
screen "Root screen" 800x480, template "Main"
   Rectangle "Rectangle_1" at 7,7 size 265x142
      Appearance <- "Comm_1_DB_Warning"
   GraphicView "Graphic view_4" at 169,29 size 84x118; Picture "h2o_1"
   GraphicView "Graphic view_2" at 89,29 size 84x118; Picture "h2o_1"
   Bar "Bar_1" at 229,7 size 43x142; Unit %; MinimumValue 0; MaximumValue 100
      ProcessValue <- "Comm_1_DB_Level"
   GraphicView "Graphic view_1" at 9,29 size 84x118; Picture "h2o_1"
   GraphicIOField "Graphic I/O field_7" at 101,119 size 76x24; PictureList "L_1"
      ProcessValue <- "Comm_1_DB_Mix_2_Status"
   GraphicIOField "Graphic I/O field_8" at 191,119 size 76x24; PictureList "L_1"
      ProcessValue <- "Comm_1_DB_Mix_3_Status"
   GraphicIOField "Graphic I/O field_6" at 12,119 size 76x24; PictureList "L_1"
      ProcessValue <- "Comm_1_DB_Mix_1_Status"
   TextField "Text field_4" at 447,6 size 223x27; Text 'мастер шкаф дозации'
   TextField "Text field_5" at 447,27 size 227x72; Text 'PolyMix'
   Button "Button_8" at 543,238 size 175x60; TextOff 'Авто'
      on Click: SetBit("Logick_DB_Start")
      Appearance <- "Logick_DB_Start"
   Button "Button_9" at 543,326 size 175x60; TextOff 'Стоп'
      on Click: ResetBit("Logick_DB_Start")
   Button "Button_10" at 543,415 size 175x60; TextOff 'Ручной'; Authorization "Operator"
      on Click: InvertBit("Logick_DB_Hand")
      Appearance <- "Logick_DB_Hand"
   Group "Group" at 7,7 size 265x142; Picture "h2o_1"; PictureList "L_1"
   Group "Group_1" at 7,160 size 265x142; Picture "h2o_1"; PictureList "L_1"
   GraphicIOField "Graphic I/O field_4" at 7,312 size 90x90; PictureList "Pump"
      ProcessValue <- "Motors_DB_M1_Status"
   GraphicIOField "Graphic I/O field_5" at 221,312 size 90x90; PictureList "Pump"
      ProcessValue <- "Motors_DB_M2_Status"
   GraphicIOField "Graphic I/O field_9" at 439,312 size 90x90; PictureList "Pump"
      ProcessValue <- "Motors_DB_M3_Status"
   Button "Button_7" at 7,402 size 90x22; TextOff 'Активен'; TextList "Hand"
      on Click: InvertBit("Logick_DB_Use_M1")
      ProcessValue <- "Motors_DB_M1_CMD_Hand"
      Appearance <- "Logick_DB_Use_M1"
   Button "Button_1" at 439,402 size 90x22; TextOff 'Активен'; TextList "Hand"
      on Click: InvertBit("Logick_DB_Use_M3")
      ProcessValue <- "Motors_DB_M1_CMD_Hand"
      Appearance <- "Logick_DB_Use_M3"
   Button "Button_2" at 221,402 size 90x22; TextOff 'Резерв М1'; TextList "Hand"
      on Click: SetBit("Logick_DB_Res_M1"); ResetBit("Logick_DB_Res_M3")
      ProcessValue <- "Motors_DB_M1_CMD_Hand"
      Appearance <- "Logick_DB_Res_M1"
   Button "Button_3" at 221,429 size 90x22; TextOff 'Резерв М3'; TextList "Hand"
      on Click: SetBit("Logick_DB_Res_M3"); ResetBit("Logick_DB_Res_M1")
      ProcessValue <- "Motors_DB_M1_CMD_Hand"
      Appearance <- "Logick_DB_Res_M3"
   Button "Button_4" at 221,457 size 90x22; TextOff 'Стоп'; TextList "Hand"
      on Click: ResetBit("Logick_DB_Res_M3"); ResetBit("Logick_DB_Res_M1")
      ProcessValue <- "Motors_DB_M1_CMD_Hand"
   GraphicView "Graphic view_7" at 275,7 size 156x149; Picture "Graphic_9"
   GraphicView "Graphic view_8" at 276,160 size 156x149; Picture "Graphic_9"
   IOField "I/O field_17" at 308,18 size 98x30; FormatPattern 99999.99
      ProcessValue <- "Statistics_DB_Mass_1"
      Appearance <- "DIx_DB_Mass_1_Signal"
   TextField "Text field_1" at 345,43 size 25x27; Text 'кг'
   IOField "I/O field_1" at 308,109 size 98x30; FormatPattern 99999.99
      ProcessValue <- "Statistics_DB_Today_1"
      Appearance <- "DIx_DB_Mass_1_Signal"
   TextField "Text field_2" at 315,83 size 85x27; Text 'за день:'
   IOField "I/O field_2" at 308,171 size 98x30; FormatPattern 99999.99
      ProcessValue <- "Statistics_DB_Mass_2"
      Appearance <- "DIx_DB_Mass_2_Signal"
   TextField "Text field_3" at 345,196 size 25x27; Text 'кг'
   IOField "I/O field_3" at 308,262 size 98x30; FormatPattern 99999.99
      ProcessValue <- "Statistics_DB_Today_2"
      Appearance <- "DIx_DB_Mass_2_Signal"
   TextField "Text field_6" at 315,236 size 85x27; Text 'за день:'
   IOField "I/O field_4" at 7,432 size 92x30; FormatPattern 9999.99
      Appearance <- "Logick_DB_Low_REQ"
      ProcessValue <- "AIx_DB_Flow_1_Result"
   TextField "Text field_7" at 33,453 size 40x27; Text 'л/ч'
   IOField "I/O field_5" at 438,432 size 92x30; FormatPattern 9999.99
      Appearance <- "Logick_DB_Low_REQ"
      ProcessValue <- "AIx_DB_Flow_2_Result"
   TextField "Text field_8" at 464,453 size 40x27; Text 'л/ч'
   Button "Button_5" at 128,362 size 60x60; TextOff 'Text'; PictureOff "table"
      on Click: ActivateScreen("Point_1", 0)
   Button "Button_6" at 348,362 size 60x60; TextOff 'Text'; PictureOff "table"
      on Click: ActivateScreen("Point_2", 0)
   TextField "Text field_9" at 347,304 size 60x27; Text 'Доза:'
   TextField "Text field_11" at 32,339 size 34x27; Text 'М1'
   TextField "Text field_12" at 247,338 size 34x27; Text 'М2'
   TextField "Text field_13" at 465,337 size 34x27; Text 'М3'
   IOField "I/O field_7" at 119,328 size 77x30; FormatPattern 999.99
      ProcessValue <- "Logick_DB_D_1"
      Visibility <- "Logick_DB_Fix_1"
   TextField "Text field_14" at 128,303 size 60x27; Text 'Доза:'
   Button "Button_12" at 118,424 size 80x25; TextOff 'Text'; Authorization "Operator"; PictureList "ON_OFF"
      on Click: InvertBit("Logick_DB_Fix_1")
      ProcessValue <- "Logick_DB_Fix_1"
   IOField "I/O field_8" at 119,328 size 77x30; Authorization "Operator"; FormatPattern 999.99
      ProcessValue <- "Logick_DB_Fix_D_1"
      Visibility <- "Logick_DB_Fix_1"
   IOField "I/O field_6" at 339,329 size 77x30; FormatPattern 999.99
      Visibility <- "Logick_DB_Fix_2"
      ProcessValue <- "Logick_DB_D_2"
   Button "Button_11" at 339,424 size 80x25; TextOff 'Text'; PictureList "ON_OFF"; Authorization "Operator"
      on Click: InvertBit("Logick_DB_Fix_2")
      ProcessValue <- "Logick_DB_Fix_2"
   IOField "I/O field_9" at 339,329 size 77x30; Authorization "Operator"; FormatPattern 999.99
      Visibility <- "Logick_DB_Fix_2"
      ProcessValue <- "Logick_DB_Fix_D_2"
   Button "Button_13" at 8,312 size 86x86; TextOff 'Text'
      on Click: InvertBit("Motors_DB_M1_CMD_Start_M")
   Button "Button_14" at 223,312 size 86x86; TextOff 'Text'
      on Click: InvertBit("Motors_DB_M2_CMD_Start_M")
   Button "Button_15" at 441,312 size 86x86; TextOff 'Text'
      on Click: InvertBit("Motors_DB_M3_CMD_Start_M")
   TextField "Text field_16" at 447,99 size 220x27; Text 'Производительность:'
   TextField "Text field_17" at 447,127 size 112x27; Text 'Дозатор 1:'
   TextField "Text field_18" at 447,163 size 112x27; Text 'Дозатор 2:'
   TextField "Text field_19" at 447,200 size 112x27; Text 'Дозатор 3:'
   IOField "I/O field_10" at 558,127 size 77x30; Authorization "Operator"; FormatPattern 9999
      ProcessValue <- "AOx_DB_M1_SP_SP_M"
      Appearance <- "AOx_DB_M1_SP_CMD_Hand"
   IOField "I/O field_11" at 558,162 size 77x30; Authorization "Operator"; FormatPattern 9999
      Appearance <- "AOx_DB_M2_SP_CMD_Hand"
      ProcessValue <- "AOx_DB_M2_SP_SP_M"
   IOField "I/O field_12" at 558,197 size 77x30; Authorization "Operator"; FormatPattern 9999
      Appearance <- "AOx_DB_M3_SP_CMD_Hand"
      ProcessValue <- "AOx_DB_M3_SP_SP_M"
   IOField "I/O field_13" at 339,448 size 80x30; FormatPattern 999.99
      ProcessValue <- "AIx_DB_Trans_2_Result"
   IOField "I/O field_14" at 118,448 size 80x30; FormatPattern 999.99
      ProcessValue <- "AIx_DB_Trans_1_Result"
   Button "Button_16" at 278,6 size 149x139; TextOff 'Text'
      on Click: ActivateScreen("Mass_1", 0)
   Button "Button_17" at 280,159 size 149x139; TextOff 'Text'
      on Click: ActivateScreen("Mass_2", 0)
   GraphicView "Graphic view_9" at 447,236 size 30x30; Picture "heat"
      Appearance <- "DIx_DB_Heat_1_Signal"
   GraphicView "Graphic view_10" at 492,236 size 30x30; Picture "heat"
      Appearance <- "DIx_DB_Heat_2_Signal"
   GraphicView "Graphic view_11" at 448,274 size 30x30; Picture "heat"
      Appearance <- "DIx_DB_Heat_3_Signal"
   GraphicView "Graphic view_12" at 492,274 size 30x30; Picture "heat"
      Appearance <- "DIx_DB_Heat_4_Signal"
   IOField "I/O field_19" at 637,127 size 92x30; FormatPattern 9999.99
      Appearance <- "Logick_DB_Low_REQ"
      ProcessValue <- "AIx_DB_Flow_3_Result"
   IOField "I/O field_16" at 637,197 size 92x30; FormatPattern 9999.99
      Appearance <- "Logick_DB_Low_REQ"
      ProcessValue <- "AIx_DB_Flow_4_Result"
   TextField "Text field_22" at 663,164 size 40x27; Text 'л/ч'
   Rectangle "Rectangle_8" at 36,90 size 175x115
      Visibility <- "Any_Hand"
      Appearance <- "Any_Hand"
   TextField "Text field_10" at 40,97 size 169x99; Text 'Внимание! Часть устройств в ручном режиме. Корректная работа невозможна.'
      Visibility <- "Any_Hand"
      Appearance <- "Any_Hand"
   Button "Button_19" at 151,351 size 150x32; TextOff 'Игнорировать'
      on Click: SetBit("Logick_DB_Low_CMD")
      Visibility <- "Logick_DB_Low_view"
      Appearance <- "Logick_DB_Low_CMD"
   Rectangle "Rectangle_12" at 19,257 size 406x145
      Visibility <- "Logick_DB_Low_view"
   TextField "Text field_15" at 324,302 size 19x27; Text 'м'
      Visibility <- "Logick_DB_Low_view"
   IOField "I/O field_15" at 286,301 size 37x32; FormatPattern 99
      Visibility <- "Logick_DB_Low_view"
      ProcessValue <- "Logick_DB_Low_SP_M"
   TextField "Text field_20" at 107,301 size 175x27; Text 'остановка через:'
      Visibility <- "Logick_DB_Low_view"
   TextField "Text field_21" at 108,271 size 234x27; Text 'Низая уставка дозации'
      Visibility <- "Logick_DB_Low_view"
   Button "Button_18" at 151,350 size 150x32; TextOff 'Игнорировать'
      on Click: SetBit("Logick_DB_Low_CMD")
      Visibility <- "Logick_DB_Low_view"
      Appearance <- "Logick_DB_Low_CMD"
   Rectangle "Rectangle_3" at 7,160 size 265x142
      Appearance <- "Comm_2_DB_Warning"
   GraphicView "Graphic view_3" at 169,182 size 84x118; Picture "h2o_1"
   GraphicView "Graphic view_5" at 89,182 size 84x118; Picture "h2o_1"
   Bar "Bar_2" at 229,160 size 43x142; Unit %; MinimumValue 0; MaximumValue 100
      ProcessValue <- "Comm_2_DB_Level"
   GraphicView "Graphic view_6" at 9,182 size 84x118; Picture "h2o_1"
   GraphicIOField "Graphic I/O field_1" at 101,272 size 76x24; PictureList "L_1"
      ProcessValue <- "Comm_2_DB_Mix_2_Status"
   GraphicIOField "Graphic I/O field_2" at 191,272 size 76x24; PictureList "L_1"
      ProcessValue <- "Comm_2_DB_Mix_3_Status"
   GraphicIOField "Graphic I/O field_3" at 12,272 size 76x24; PictureList "L_1"
      ProcessValue <- "Comm_2_DB_Mix_1_Status"

screen "Alarms" 800x480, template "Main"
   AlarmView "Alarm view_1" at 4,3 size 718x470; ColumnTextDate 'Дата'; ColumnTextAlarmState 'Статус'; ColumnTextTime 'Время'; ColumnTextAlarmText 'Аварийное сообщение'

screen "SIMATIC PLC system diagnostics" 800x480, template "Main"
   SysDiagControl "HmiScreenItemData" at 1,49 size 796x423
   Button "Back" at 1,1 size 159x47; TextOn 'Back'; TextOff 'Back'
      on Release: ActivateScreen("System screens", 0)

screen "System information" 800x480, template "Main"
   TextField "HmiScreenItemData" at 35,51 size 171x28; Text 'HMI device type:'
   TextField "HmiScreenItemData_1" at 241,51 size 524x28; Text 'KTP700 Basic+ PN 14.0.1.0'
   TextField "HmiScreenItemData_2" at 35,81 size 171x28; Text 'Connection:'
   TextField "HmiScreenItemData_3" at 241,81 size 524x28; Text 'PROFINET (X1)'
   TextField "HmiScreenItemData_4" at 35,111 size 171x28; Text 'PLC:'
   TextField "HmiScreenItemData_5" at 241,111 size 524x28; Text 'SIMATIC S7 1200'
   Button "Back" at 1,1 size 159x47; TextOn 'Back'; TextOff 'Back'
      on Release: ActivateScreen("System screens", 0)

screen "System screens" 800x480, template "Main"
   Button "Back" at 1,1 size 159x47; TextOn 'Back'; TextOff 'Back'
      on Release: ActivateScreen("Root screen", 0)
   Button "HmiScreenItemData" at 36,95 size 159x47; TextOn 'SIMATIC PLC system diagnos...'; TextOff 'SIMATIC PLC system diagnos...'; PictureOn "Navigates to SIMATIC PLC system diagnostics for KTP700 Basic+ PN 14.0.1.0"; PictureOff "Navigates to SIMATIC PLC system diagnostics for KTP700 Basic+ PN 14.0.1.0"
      on Release: ActivateScreen("SIMATIC PLC system diagnostics", 0)
   Button "HmiScreenItemData_1" at 36,154 size 159x47; TextOn 'Project information'; TextOff 'Project information'; PictureOn "Navigates to Project information for KTP700 Basic+ PN 14.0.1.0"; PictureOff "Navigates to Project information for KTP700 Basic+ PN 14.0.1.0"
      on Release: ActivateScreen("Project information", 0)
   Button "HmiScreenItemData_2" at 36,213 size 159x47; TextOn 'System information'; TextOff 'System information'; PictureOn "Navigates to System information for KTP700 Basic+ PN 14.0.1.0"; PictureOff "Navigates to System information for KTP700 Basic+ PN 14.0.1.0"
      on Release: ActivateScreen("System information", 0)
   Button "HmiScreenItemData_3" at 36,272 size 159x47; TextOn 'Different jobs'; TextOff 'Different jobs'; PictureOn "Navigates to Different jobs for KTP700 Basic+ PN 14.0.1.0"; PictureOff "Navigates to Different jobs for KTP700 Basic+ PN 14.0.1.0"
      on Release: ActivateScreen("Different jobs", 0)

screen "Different jobs" 800x480, template "Main"
   Button "Online" at 36,95 size 159x47; TextOn 'Online'; TextOff 'Online'
      on Release: function_bb44b551(0)
   Button "Offline" at 36,154 size 159x47; TextOn 'Offline'; TextOff 'Offline'
      on Release: function_bb44b551(1)
   Button "Transfer" at 36,213 size 159x47; TextOn 'Transfer'; TextOff 'Transfer'
      on Release: function_bb44b551(2)
   Button "Toggle language" at 36,272 size 159x47; TextOn 'Toggle language'; TextOff 'Toggle language'
      on Release: function_fb9197e8(-1)
   Button "Stop Runtime" at 36,331 size 159x47; TextOn 'Stop Runtime'; TextOff 'Stop Runtime'
      on Release: StopRuntime(0)
   Button "Back" at 1,1 size 159x47; TextOn 'Back'; TextOff 'Back'
      on Release: ActivateScreen("System screens", 0)

screen "Project information" 800x480, template "Main"
   TextField "HmiScreenItemData" at 35,51 size 171x28; Text 'Project name:'
   TextField "HmiScreenItemData_1" at 241,51 size 524x28; Text 'PolyMix_v0.1'
   TextField "HmiScreenItemData_2" at 35,81 size 171x28; Text 'Created on:'
   TextField "HmiScreenItemData_3" at 241,81 size 524x28; Text '10/24/2017 3:17:12 PM'
   TextField "HmiScreenItemData_4" at 35,111 size 171x28; Text 'Author:'
   TextField "HmiScreenItemData_5" at 241,111 size 524x28; Text 'WinCC'
   TextField "HmiScreenItemData_6" at 35,141 size 171x28; Text 'Description:'
   TextField "HmiScreenItemData_7" at 241,141 size 524x28; Text '(not configured)'
   Button "Back" at 1,1 size 159x47; TextOn 'Back'; TextOff 'Back'
      on Release: ActivateScreen("System screens", 0)

screen "SP" 800x480, template "Main"
   GraphicView "Graphic view_1" at 20,61 size 347x209; Picture "clean2"
   TextField "Text field_1" at 288,5 size 156x47; Text 'Уставки'
   TextField "Text field_2" at 129,75 size 130x33; Text 'Дозатор 1'
   TextField "Text field_12" at 28,137 size 34x23; Text 'С ='
   TextField "Text field_13" at 151,138 size 67x23; Text '% масс'
   GraphicView "Graphic view_2" at 83,133 size 66x33; Picture "input_1"
   IOField "I/O field_1" at 87,136 size 58x27; Authorization "Operator"; FormatPattern 99.99
      ProcessValue <- "Logick_DB_C_1"
   TextField "Text field_3" at 95,118 size 43x17; Text 'макс 1'
   TextField "Text field_4" at 90,163 size 53x17; Text 'мин 0.05'
   TextField "Text field_5" at 30,188 size 45x23; Text 'Доза'
   IOField "I/O field_7" at 84,188 size 65x27; FormatPattern 999.99
      Visibility <- "Logick_DB_Fix_1"
      ProcessValue <- "Logick_DB_D_1"
   GraphicView "Graphic view_3" at 80,185 size 73x33; Picture "input_1"
   IOField "I/O field_8" at 84,188 size 65x27; Authorization "Operator"; FormatPattern 999.99
      ProcessValue <- "Logick_DB_Fix_D_1"
   Button "Button_12" at 161,227 size 80x25; TextOff 'Text'; PictureList "ON_OFF"; Authorization "Operator"
      on Click: InvertBit("Logick_DB_Fix_1")
      ProcessValue <- "Logick_DB_Fix_1"
   TextField "Text field_6" at 33,226 size 126x23; Text 'Фиксированно'
   Button "Button_5" at 288,192 size 60x60; TextOff 'Text'; PictureOff "table"
      on Click: ActivateScreen("Point_1", 0)
   GraphicView "Graphic view_4" at 374,61 size 347x209; Picture "clean2"
   TextField "Text field_7" at 483,75 size 130x33; Text 'Дозатор 2'
   TextField "Text field_8" at 382,137 size 34x23; Text 'С ='
   TextField "Text field_9" at 505,138 size 67x23; Text '% масс'
   GraphicView "Graphic view_5" at 437,133 size 66x33; Picture "input_1"
   IOField "I/O field_2" at 441,136 size 58x27; Authorization "Operator"; FormatPattern 99.99
      ProcessValue <- "Logick_DB_C_2"
   TextField "Text field_10" at 449,118 size 43x17; Text 'макс 1'
   TextField "Text field_11" at 444,163 size 53x17; Text 'мин 0.05'
   TextField "Text field_14" at 384,188 size 45x23; Text 'Доза'
   IOField "I/O field_3" at 438,188 size 65x27; FormatPattern 999.99
      ProcessValue <- "Logick_DB_D_2"
      Visibility <- "Logick_DB_Fix_2"
   GraphicView "Graphic view_6" at 434,185 size 73x33; Picture "input_1"
   IOField "I/O field_4" at 438,188 size 65x27; Authorization "Operator"; FormatPattern 999.99
      ProcessValue <- "Logick_DB_Fix_D_2"
   Button "Button_1" at 515,227 size 80x25; TextOff 'Text'; Authorization "Operator"; PictureList "ON_OFF"
      on Click: InvertBit("Logick_DB_Fix_2")
      ProcessValue <- "Logick_DB_Fix_2"
   TextField "Text field_15" at 387,226 size 126x23; Text 'Фиксированно'
   Button "Button_2" at 642,192 size 60x60; TextOff 'Text'; PictureOff "table"
      on Click: ActivateScreen("Point_2", 0)
   GraphicView "Graphic view_7" at 20,270 size 347x209; Picture "clean2"
   TextField "Text field_16" at 108,284 size 172x33; Text 'Ограничения'
   TextField "Text field_17" at 29,341 size 201x23; Text 'Макс уставка дозатора'
   IOField "I/O field_5" at 241,341 size 65x27; FormatPattern 999.99
      ProcessValue <- "Logick_DB_D_1"
      Visibility <- "Logick_DB_Fix_1"
   GraphicView "Graphic view_8" at 237,338 size 73x33; Picture "input_1"
   IOField "I/O field_6" at 241,341 size 65x27; Authorization "Operator"; FormatPattern 9999
      ProcessValue <- "Logick_DB_Max_SP"
   TextField "Text field_18" at 309,341 size 34x23; Text 'л/ч'
   TextField "Text field_19" at 29,378 size 193x23; Text 'Мин уставка дозатора'
   IOField "I/O field_9" at 241,378 size 65x27; FormatPattern 999.99
      Visibility <- "Logick_DB_Fix_1"
      ProcessValue <- "Logick_DB_D_1"
   GraphicView "Graphic view_9" at 237,375 size 73x33; Picture "input_1"
   IOField "I/O field_10" at 241,378 size 65x27; Authorization "Operator"; FormatPattern 9999
      ProcessValue <- "Logick_DB_Min_SP"
   TextField "Text field_20" at 309,378 size 34x23; Text 'л/ч'
   TextField "Text field_21" at 29,415 size 166x23; Text 'Время до останова'
   IOField "I/O field_11" at 241,415 size 65x27; FormatPattern 999.99
      ProcessValue <- "Logick_DB_D_1"
      Visibility <- "Logick_DB_Fix_1"
   GraphicView "Graphic view_10" at 237,412 size 73x33; Picture "input_1"
   IOField "I/O field_12" at 241,415 size 65x27; Authorization "Operator"; FormatPattern 9999
      ProcessValue <- "Logick_DB_Low_SP_M"
   TextField "Text field_22" at 309,415 size 17x23; Text 'м'
   TextField "Text field_23" at 29,444 size 94x23; Text 'Остановка'
   Button "Button_3" at 147,443 size 80x25; TextOff 'Text'; PictureList "ON_OFF"; Authorization "Operator"
      on Click: InvertBit("Logick_DB_Low_use")
      ProcessValue <- "Logick_DB_Low_use"
   Button "HmiScreenItemData_4" at 374,271 size 347x47; TextOn 'О нас'; TextOff 'Статистика весов 1'; PictureOn "Navigates to System screens for KTP700 Basic+ PN 14.0.1.0"; PictureOff "Navigates to System screens for KTP700 Basic+ PN 14.0.1.0"
      on Release: ActivateScreen("Mass_1", 0)
   Button "HmiScreenItemData_1" at 374,323 size 347x47; TextOn 'О нас'; TextOff 'Статистика весов 2'; PictureOn "Navigates to System screens for KTP700 Basic+ PN 14.0.1.0"; PictureOff "Navigates to System screens for KTP700 Basic+ PN 14.0.1.0"
      on Release: ActivateScreen("Mass_2", 0)
   Button "Button_4" at 559,382 size 80x25; TextOff 'Text'; PictureList "ON_OFF"; Authorization "Operator"
      on Click: InvertBit("Logick_DB_Correction_1")
      ProcessValue <- "Logick_DB_Correction_1"
   TextField "Text field_24" at 375,381 size 179x23; Text 'Коррекция насоса 1:'
   Button "Button_6" at 559,404 size 80x25; TextOff 'Text'; Authorization "Operator"; PictureList "ON_OFF"
      on Click: InvertBit("Logick_DB_Correction_2")
      ProcessValue <- "Logick_DB_Correction_2"
   TextField "Text field_25" at 375,403 size 179x23; Text 'Коррекция насоса 2:'
   IOField "I/O field_13" at 652,384 size 65x21; Authorization "Operator"; FormatPattern 9.99
      ProcessValue <- "Logick_DB_C_SP_1"
   IOField "I/O field_15" at 652,406 size 65x21; Authorization "Operator"; FormatPattern 9.99
      ProcessValue <- "Logick_DB_C_SP_2"

screen "Wieght" 800x480, template "Main"
   GraphicView "Graphic view_1" at 20,61 size 347x209; Picture "clean2"
   TextField "Text field_1" at 256,5 size 233x47; Text 'Калибровка'
   TextField "Text field_2" at 149,75 size 90x33; Text 'Весы 1'
   TextField "Text field_6" at 268,130 size 23x23; Text 'кг'
   TextField "Text field_7" at 28,131 size 154x23; Text 'Показания весов:'
   GraphicView "Graphic view_4" at 180,126 size 89x33; Picture "input_1"
   IOField "I/O field_8" at 185,129 size 80x27; Authorization "Operator"; FormatPattern 999999.9
      ProcessValue <- "RS232_DB_Mass_1"
   GraphicView "Graphic view_5" at 374,61 size 347x209; Picture "clean2"
   TextField "Text field_21" at 503,75 size 90x33; Text 'Весы 2'
   TextField "Text field_3" at 267,172 size 23x23; Text 'кг'
   TextField "Text field_4" at 27,173 size 87x23; Text 'Вес тары:'
   GraphicView "Graphic view_2" at 179,168 size 89x33; Picture "input_1"
   IOField "I/O field_1" at 184,171 size 80x27; Authorization "Operator"; FormatPattern 999999.9
      ProcessValue <- "Statistics_DB_Zero_1"
   TextField "Text field_5" at 266,213 size 23x23; Text 'кг'
   TextField "Text field_8" at 26,214 size 145x23; Text 'Масса продукта:'
   GraphicView "Graphic view_3" at 178,209 size 89x33; Picture "input_1"
   IOField "I/O field_2" at 183,212 size 80x27; Authorization "Operator"; FormatPattern 999999.9
      ProcessValue <- "Statistics_DB_Mass_1"
   TextField "Text field_9" at 624,128 size 23x23; Text 'кг'
   TextField "Text field_10" at 384,129 size 154x23; Text 'Показания весов:'
   GraphicView "Graphic view_6" at 536,124 size 89x33; Picture "input_1"
   IOField "I/O field_3" at 541,127 size 80x27; Authorization "Operator"; FormatPattern 999999.9
      ProcessValue <- "RS232_DB_Mass_2"
   TextField "Text field_11" at 623,170 size 23x23; Text 'кг'
   TextField "Text field_12" at 383,171 size 87x23; Text 'Вес тары:'
   GraphicView "Graphic view_7" at 535,166 size 89x33; Picture "input_1"
   IOField "I/O field_4" at 540,169 size 80x27; Authorization "Operator"; FormatPattern 999999.9
      ProcessValue <- "Statistics_DB_Zero_2"
   TextField "Text field_13" at 622,211 size 23x23; Text 'кг'
   TextField "Text field_14" at 382,212 size 145x23; Text 'Масса продукта:'
   GraphicView "Graphic view_8" at 534,207 size 89x33; Picture "input_1"
   IOField "I/O field_5" at 539,210 size 80x27; Authorization "Operator"; FormatPattern 999999.9
      ProcessValue <- "Statistics_DB_Mass_2"
   GraphicView "Graphic view_9" at 20,271 size 347x209; Picture "clean2"
   TextField "Text field_15" at 120,286 size 148x33; Text 'Учёт веса 1'
   GraphicView "Graphic view_10" at 372,270 size 347x209; Picture "clean2"
   TextField "Text field_16" at 474,284 size 148x33; Text 'Учёт веса 2'
   TextField "Text field_17" at 32,331 size 81x23; Text 'Текущий'
   TextField "Text field_18" at 32,359 size 85x23; Text 'Прошлый'
   TextField "Text field_19" at 32,387 size 110x23; Text 'Дельта макс'
   TextField "Text field_20" at 32,415 size 102x23; Text 'Дельта мин'
   TextField "Text field_22" at 32,439 size 153x23; Text 'Время измерения'
   TextField "Text field_23" at 296,337 size 23x23; Text 'кг'
   GraphicView "Graphic view_11" at 208,333 size 89x26; Picture "input_1"
   IOField "I/O field_6" at 213,336 size 80x19; Authorization "Operator"; FormatPattern 999999.9
      ProcessValue <- "Statistics_DB_Mass_1"
   TextField "Text field_24" at 295,363 size 23x23; Text 'кг'
   GraphicView "Graphic view_12" at 207,359 size 89x26; Picture "input_1"
   IOField "I/O field_7" at 212,362 size 80x19; Authorization "Operator"; FormatPattern 999999.9
      ProcessValue <- "Statistics_DB_Last_1"
   TextField "Text field_25" at 295,389 size 23x23; Text 'кг'
   GraphicView "Graphic view_13" at 207,385 size 89x26; Picture "input_1"
   IOField "I/O field_9" at 212,388 size 80x19; Authorization "Developer"; FormatPattern 999999.9
      ProcessValue <- "Statistics_DB_Max_D_1"
   TextField "Text field_26" at 294,415 size 23x23; Text 'кг'
   GraphicView "Graphic view_14" at 206,411 size 89x26; Picture "input_1"
   IOField "I/O field_10" at 212,414 size 80x19; Authorization "Developer"; FormatPattern 999999.9
      ProcessValue <- "Statistics_DB_Min_D_1"
   TextField "Text field_27" at 243,440 size 17x23; Text 'м'
   GraphicView "Graphic view_15" at 209,437 size 36x26; Picture "input_1"
   IOField "I/O field_11" at 212,440 size 31x19; Authorization "Developer"; FormatPattern 999
      ProcessValue <- "Statistics_DB_T_SP_M"
   GraphicView "Graphic view_16" at 123,346 size 89x26; Picture "input_1"
   IOField "I/O field_12" at 128,349 size 80x19; Authorization "Operator"; FormatPattern 999999.9
      ProcessValue <- "Statistics_DB_Delta_1"
   TextField "Text field_28" at 294,440 size 13x23; Text 'с'
   GraphicView "Graphic view_17" at 259,437 size 36x26; Picture "input_1"
   IOField "I/O field_13" at 261,440 size 31x19; Authorization "Developer"; FormatPattern 99
      ProcessValue <- "Statistics_DB_T_SP_S"
   Button "Button_1" at 25,273 size 110x19; TextOff 'Синхронизировать'
      on Click: SetBit("Sync")
   Button "Button_2" at 377,272 size 110x19; TextOff 'Синхронизировать'
      on Click: SetBit("Sync_2")
   TextField "Text field_29" at 380,335 size 81x23; Text 'Текущий'
   TextField "Text field_30" at 380,363 size 85x23; Text 'Прошлый'
   TextField "Text field_31" at 380,391 size 110x23; Text 'Дельта макс'
   TextField "Text field_32" at 380,419 size 102x23; Text 'Дельта мин'
   TextField "Text field_33" at 380,443 size 153x23; Text 'Время измерения'
   TextField "Text field_34" at 644,341 size 23x23; Text 'кг'
   GraphicView "Graphic view_18" at 556,337 size 89x26; Picture "input_1"
   IOField "I/O field_14" at 561,340 size 80x19; Authorization "Operator"; FormatPattern 999999.9
      ProcessValue <- "Statistics_DB_Mass_2"
   TextField "Text field_35" at 643,367 size 23x23; Text 'кг'
   GraphicView "Graphic view_19" at 555,363 size 89x26; Picture "input_1"
   IOField "I/O field_15" at 560,366 size 80x19; Authorization "Operator"; FormatPattern 999999.9
      ProcessValue <- "Statistics_DB_Last_2"
   TextField "Text field_36" at 643,393 size 23x23; Text 'кг'
   GraphicView "Graphic view_20" at 555,389 size 89x26; Picture "input_1"
   IOField "I/O field_16" at 560,392 size 80x19; Authorization "Developer"; FormatPattern 999999.9
      ProcessValue <- "Statistics_DB_Max_D_2"
   TextField "Text field_37" at 642,419 size 23x23; Text 'кг'
   GraphicView "Graphic view_21" at 554,415 size 89x26; Picture "input_1"
   IOField "I/O field_17" at 560,418 size 80x19; Authorization "Developer"; FormatPattern 999999.9
      ProcessValue <- "Statistics_DB_Min_D_2"
   TextField "Text field_38" at 591,444 size 17x23; Text 'м'
   GraphicView "Graphic view_22" at 557,441 size 36x26; Picture "input_1"
   IOField "I/O field_18" at 560,444 size 31x19; Authorization "Developer"; FormatPattern 999
      ProcessValue <- "Statistics_DB_T_SP_M"
   GraphicView "Graphic view_23" at 471,350 size 89x26; Picture "input_1"
   IOField "I/O field_19" at 476,353 size 80x19; Authorization "Operator"; FormatPattern 999999.9
      ProcessValue <- "Statistics_DB_Delta_2"
   TextField "Text field_39" at 642,444 size 13x23; Text 'с'
   GraphicView "Graphic view_24" at 607,441 size 36x26; Picture "input_1"
   IOField "I/O field_20" at 609,444 size 31x19; Authorization "Developer"; FormatPattern 99
      ProcessValue <- "Statistics_DB_T_SP_S"

screen "Monitor" 800x480, template "Main"
   Button "HmiScreenItemData_1" at 10,425 size 159x47; TextOff 'Система'; PictureOn "Navigates to System screens for KTP700 Basic+ PN 14.0.1.0"; PictureOff "Navigates to System screens for KTP700 Basic+ PN 14.0.1.0"; Authorization "Admin"
      on Release: ActivateScreen("System screens", 0)
   Button "HmiScreenItemData_3" at 380,425 size 159x47; TextOff 'Настройки'; PictureOn "Navigates to System screens for KTP700 Basic+ PN 14.0.1.0"; PictureOff "Navigates to System screens for KTP700 Basic+ PN 14.0.1.0"; Authorization "Admin"
      on Release: ActivateScreen("Settings", 0); SetTag("settings", 0)
   Button "HmiScreenItemData_4" at 565,425 size 159x47; TextOn 'О нас'; TextOff 'О нас'; PictureOn "Navigates to System screens for KTP700 Basic+ PN 14.0.1.0"; PictureOff "Navigates to System screens for KTP700 Basic+ PN 14.0.1.0"
      on Release: ActivateScreen("About", 0)
   TextField "Text field_1" at 168,4 size 424x47; Text 'Параметры установки'
   TextField "Text field_2" at 261,56 size 262x33; Text 'Состояние сигналов'
   TextField "Text field_3" at 71,92 size 189x27; Text 'Дискретные входа'
   TextField "Text field_4" at 477,92 size 205x27; Text 'Дискретные выхода'
   TextField "Text field_5" at 282,340 size 189x27; Text 'Аналоговые входа'
   TextField "Text field_6" at 43,117 size 254x23; Text 'I 0.0 - Дозатор 1 - Готовность'
   TextField "Text field_7" at 43,138 size 254x23; Text 'I 0.1 - Дозатор 2 - Готовность'
   TextField "Text field_8" at 43,160 size 254x23; Text 'I 0.2 - Дозатор 3 - Готовность'
   TextField "Text field_9" at 43,181 size 274x23; Text 'I 0.3 - Нагреватель 1 - В работе'
   TextField "Text field_10" at 43,203 size 274x23; Text 'I 0.4 - Нагреватель 2 - В работе'
   TextField "Text field_11" at 43,224 size 274x23; Text 'I 0.5 - Нагреватель 3 - В работе'
   TextField "Text field_12" at 43,246 size 274x23; Text 'I 0.6 - Нагреватель 4 - В работе'
   TextField "Text field_13" at 43,267 size 207x23; Text 'I 0.7 - Внешний останов'
   TextField "Text field_14" at 43,289 size 208x23; Text 'I 1.0 - Весы 1 - В работе'
   TextField "Text field_15" at 43,310 size 208x23; Text 'I 1.1 - Весы 2 - В работе'
   Circle "Circle_1" at 10,120 size 17x17
      Appearance <- "DIx_DB_M1_QF_Signal"
   Circle "Circle_2" at 10,141 size 17x17
      Appearance <- "DIx_DB_M2_QF_Signal"
   Circle "Circle_3" at 10,163 size 17x17
      Appearance <- "DIx_DB_M3_QF_Signal"
   Circle "Circle_4" at 10,184 size 17x17
      Appearance <- "DIx_DB_Heat_1_Signal"
   Circle "Circle_5" at 10,206 size 17x17
      Appearance <- "DIx_DB_Heat_2_Signal"
   Circle "Circle_6" at 10,227 size 17x17
      Appearance <- "DIx_DB_Heat_3_Signal"
   Circle "Circle_7" at 10,249 size 17x17
      Appearance <- "DIx_DB_Heat_4_Signal"
   Circle "Circle_8" at 10,270 size 17x17
      Appearance <- "DIx_DB_AllBlock_Signal"
   Circle "Circle_9" at 10,292 size 17x17
      Appearance <- "DIx_DB_Mass_1_Signal"
   Circle "Circle_10" at 10,313 size 17x17
      Appearance <- "DIx_DB_Mass_2_Signal"
   TextField "Text field_20" at 447,117 size 222x23; Text 'Q 0.0 - Дозатор 1 - Запуск'
   TextField "Text field_21" at 447,139 size 222x23; Text 'Q 0.1 - Дозатор 2 - Запуск'
   TextField "Text field_22" at 447,160 size 222x23; Text 'Q 0.2 - Дозатор 3 - Запуск'
   TextField "Text field_23" at 447,182 size 204x23; Text 'Q 0.3 - Авария шкафа 1'
   TextField "Text field_24" at 447,203 size 204x23; Text 'Q 0.4 - Авария шкафа 2'
   TextField "Text field_25" at 447,225 size 187x23; Text 'Q 0.5 - Общая авария'
   TextField "Text field_26" at 447,246 size 224x23; Text 'Q 0.6 - Авария дозатора 1'
   TextField "Text field_27" at 447,268 size 224x23; Text 'Q 0.7 - Авария дозатора 2'
   TextField "Text field_28" at 447,289 size 224x23; Text 'Q 1.0 - Авария дозатора 3'
   Circle "Circle_15" at 414,120 size 17x17
      Appearance <- "DOx_DB_M1_CMD_Q"
   Circle "Circle_16" at 414,142 size 17x17
      Appearance <- "DOx_DB_M2_CMD_Q"
   Circle "Circle_17" at 414,163 size 17x17
      Appearance <- "DOx_DB_M3_CMD_Q"
   Circle "Circle_18" at 414,185 size 17x17
      Appearance <- "DOx_DB_LED_Error_1_Q"
   Circle "Circle_19" at 414,206 size 17x17
      Appearance <- "DOx_DB_LED_Error_2_Q"
   Circle "Circle_20" at 414,228 size 17x17
      Appearance <- "DOx_DB_LED_Alarm_Q"
   Circle "Circle_21" at 414,249 size 17x17
      Appearance <- "DOx_DB_LED_M1_Alarm_Q"
   Circle "Circle_22" at 414,271 size 17x17
      Appearance <- "DOx_DB_LED_M2_Alarm_Q"
   Circle "Circle_23" at 414,292 size 17x17
      Appearance <- "DOx_DB_LED_M3_Alarm_Q"
   TextField "Text field_30" at 414,375 size 184x23; Text 'PIW 264 - Мутность 1'
   TextField "Text field_31" at 414,398 size 184x23; Text 'PIW 266 - Мутность 2'
   IOField "I/O field_1" at 617,376 size 96x22; FormatPattern s99999
      ProcessValue <- "AIx_DB_Trans_1_Signal"
   IOField "I/O field_2" at 617,396 size 96x22; FormatPattern s99999
      ProcessValue <- "AIx_DB_Trans_2_Signal"
   TextField "Text field_16" at 9,375 size 208x23; Text 'PIW 260 - Расходомер 1'
   TextField "Text field_17" at 9,398 size 208x23; Text 'PIW 262 - Расходомер 2'
   IOField "I/O field_3" at 247,376 size 96x22; FormatPattern s99999
      ProcessValue <- "AIx_DB_Flow_1_Signal"
   IOField "I/O field_4" at 247,396 size 96x22; FormatPattern s99999
      ProcessValue <- "AIx_DB_Flow_2_Signal"

